// TIA Portal project "Mawomat" (V17)

(* hardware
DEVICE "S7-1500/ET200MP station_1"  S7-1500 station
   slot 0: "Rail_0"  Rack  6ES7 590-1***0-0AA0
   slot 1: "PLC_1"  CPU 1511-1 PN  6ES7 511-1AK00-0AB0  V1.8
      slot 3: "CPU display_1"  6ES7591-1AA00-0AA0
      slot 32768: "PROFINET interface_1"  X1
         slot 32769: "Port_1"  X1 P1
         slot 32770: "Port_2"  X1 P2
DEVICE "HMI_1"  KTP1200 Basic PN
   slot 0: "HMI_1"  KTP1200 Basic PN  6AV2 123-2MB03-0AX0  17.0.0.0
   slot 1: "HMI_RT_1"  KTP1200 Basic PN  6AV2 123-2MB03-0AX0  17.0.0.0
   slot 5: "HMI_1.IE_CP_1"  PROFINET Interface  17.0.0.0
      slot 1: "PROFINET Interface_1"  PROFINET Interface
         slot 1: "Port_1"  Port
DEVICE "SINAMICS G_1"  Sinamics.Device
   slot 0: "	_0"  Rail  SinamicsG120RackPN
   slot 0: "Drive_1"  G120 CU240E-2 PN  6SL3244-0BB12-1FA0  4.7.13
      slot 1: "PROFINET interface"  MDD-SinamicsG120-P
DEVICE "SINAMICS G_2"  Sinamics.Device
   slot 0: "	_0"  Rail  SinamicsG120RackPN
   slot 0: "Drive_2"  G120 CU240E-2 PN  6SL3244-0BB12-1FA0  4.7.13
      slot 1: "PROFINET interface"  MDD-SinamicsG120-P
*)

// ===== PLC "PLC_1"  CPU 1511-1 PN =====

VAR_GLOBAL   // PLC tag table "Default tag table"
   "System_Byte" AT %MB1 : Byte;
   "FirstScan" AT %M1.0 : Bool;
   "DiagStatusUpdate" AT %M1.1 : Bool;
   "AlwaysTRUE" AT %M1.2 : Bool;
   "AlwaysFALSE" AT %M1.3 : Bool;
   "Clock_Byte" AT %MB0 : Byte;
   "Clock_10Hz" AT %M0.0 : Bool;
   "Clock_5Hz" AT %M0.1 : Bool;
   "Clock_2.5Hz" AT %M0.2 : Bool;
   "Clock_2Hz" AT %M0.3 : Bool;
   "Clock_1.25Hz" AT %M0.4 : Bool;
   "Clock_1Hz" AT %M0.5 : Bool;
   "Clock_0.625Hz" AT %M0.6 : Bool;
   "Clock_0.5Hz" AT %M0.7 : Bool;
   "systemowe01" AT %M50.0 : Bool;
   "systemowe02" AT %M50.1 : Bool;
   "imp1s" AT %M50.2 : Bool;
   "Tag_29" AT %M51.0 : Bool;
   "Tag_28" AT %M51.1 : Bool;
   "imp0.1s" AT %M51.2 : Bool;
   "Tag_31" AT %M52.0 : Bool;
   "Tag_32" AT %M52.1 : Bool;
   "Imp0.2s" AT %M52.2 : Bool;
   "Tag_1" AT %M60.0 : Bool;
   "Tag_2" AT %M20.2 : Bool;
   "Tag_3" AT %M60.1 : Bool;
   "Tag_4" AT %M10.0 : Bool;
   "Tag_5" AT %M10.1 : Bool;
   "Tag_6" AT %M10.2 : Bool;
   "Tag_7" AT %M10.3 : Bool;
END_VAR

VAR_GLOBAL   // PLC tag table "Tag table_1"
   "qw256" AT %QW256 : Word;
END_VAR

TYPE "UDT321_DIO"
   STRUCT
      yNrPLC : Byte;   // DANE OGOLNE - Numer sterownika [0-255]
      yNrMAN : Byte;   // DANE OGOLNE - Numer powiazanej 'grupy recznej' [0-255]
      yNrID : Int;   // DANE OGOLNE - Numer ID obiektu w klasie [0-65536]
      yNrMD : Int;   // DANE OGOLNE - Numer powiazanego 'modelu drogi'
      bWeAkt : Bool;   // WEJSCIE - Aktywacja urz. w systemie (ustawiany tylko z programu)
      bWeZalAuto : Bool;   // WEJSCIE - Sterowanie urz. binarne w tr. Zdalnym-Auto: (0)- Wylacz; (1)- Zalacz
      bWeAwrZ : Bool;   // WEJSCIE - Awaria zewnetrzna: (0)-Brak; (1)-Aktywna
      bWeBlZmAuto : Bool;   // WEJŚCIE - Blokada zmiany trybu zdalnego z Auto na Man: (0)- Brak; (1)- Aktywna
      bRoZB1 : Byte := 16#5;   // !Rozkazy operetara
      bRoZB2 : Byte;   // !Rozkazy operatora - impulsy
      bSym : Word;   // !Symulacja
      bSt_Tryb : Word;   // !Stan
      bSt_Urz : Int;   // !Stan2
      bTrP : Int;   // !Tryb pracy
      bWySter : Bool;   // WYJSCIE - Sygnal zalaczenia urzadzenia
      bWyRst : Bool;   // WYJSCIE - Sygnal resetu awarii (impuls)
      yCzZadOpzZal : DWord;   // PARAMETR- Zadany czas opoznienia zalaczenia [0-255] sek.
      yCzAktOpzZal : DWord;   // PARAMETR- Aktualny czas opoznienia zalaczenia [0-255] sek.
      yCzZadOpzWyl : DWord;   // PARAMETR- Zadany czas opoznienia wylaczenia [0-255] sek.
      yCzAktOpzWyl : DWord;   // PARAMETR- Aktualny czas opoznienia wylaczenia [0-255] sek.
      bLatch : Bool;   // PARAMETR - Zatrzaskiwanie wyjscia (0) - Wylaczone; (1)-Zalaczone
      bAoff : Bool := 1;   // PARAMETR - samowylaczanie wylaczone (0); zalaczone (1)
      bHlp187 : Bool;   // WYJSCIE - Zal urz. w trybie AUTO
      bWeTrRem : Bool;
      bWeTrLok : Bool;
      bHlp186 : Bool;
      bTmr_On_Start : Bool;   // PARAMETR - Czas zadany timera filtru HH
      bTmr_Off_Start : Bool;   // PARAMETR - Czas zadany timera filtru LL
      bTmr_On_Ok : Bool;   // PARAMETR - Timer HH opoznienia zalaczenia odliczyl
      bTmr_Off_Ok : Bool;   // PARAMETR - Timer LL opoznienia zalaczenia odliczyl
   END_STRUCT;
END_TYPE

TYPE "UDT331_AI"
   STRUCT
      yNrPLC : Byte;   // DANE OGOLNE - Numer sterownika [0-255]
      yNrMAN : Byte;   // DANE OGOLNE - Numer powiazanej 'grupy recznej' [0-255]
      yNrID : Int;   // DANE OGOLNE - Numer ID obiektu w klasie [0-65536]
      yNrMD : Int;   // DANE OGOLNE - Numer powiazanego 'modelu drogi'
      bWeAkt : Bool;   // WEJSCIE - Aktywacja urz. w systemie (ustawiany tylko z programu)
      bWeAwrZ : Bool;   // WEJSCIE - Awaria zewnetrzna: (0)-Brak; (1)-Aktywna
      bWeBlZmAuto : Bool;   // WEJSCIE - Blokada zmiany trybu zdalnego z Auto na Man: (0)- Brak; (1)- Aktywna
      bWeSymUp : Bool;   // WEJSCIE - W trybie symulacji pomiaru skok w gore o rSymUp / sekunde
      bWeSymDown : Bool;   // WEJSCIE - W trybie symulacji pomiaru skok w dol o rSymDown / sekunde
      bRoZB1 : Byte := 16#01;   // !Rozkazy operetara
      bRoZB2 : Byte;   // !Rozkazy operatora - impulsy
      bSym : Word;   // !Symulacja
      bSt_Tryb : Word;   // !Stan
      bSt_Urz : Int;   // !Stan2
      bTrP : Int;   // !Tryb pracy
      bWyRst : Bool;   // WYJSCIE - Sygnal resetu awarii (impuls)
      yJednostka : Byte := 16#3;   // PARAMETR - Jednostka fizyczna
      yCzZadFiltru : Byte;   // PARAMETR - Czas zadany filtrow HH i LL [0-255] sek
      yCzasAktFiltrG : Byte := 16#3;   // PARAMETR - Czas aktualny filtru HH [0-255] sek
      yCzasAktFiltrD : Byte;   // PARAMETR - Czas aktualny filtru LL [0-255] sek
      bB : Byte;   // PARAMETR - Blokada generowania alarmow
      bAwrUst : Bool;   // PARAMETR - Reakcja na awarie toru pomiarowego: 0-na wyjsciu ZL; 1-ZH
      rZH : Real;   // PARAMETR - Zakres gorny pomiaru w jednostkach fizycznych
      rZL : Real;   // PARAMETR - Zakres dolny pomiaru w jednostkach fizycznych
      rGHH : Real;   // PARAMETR - Wartosc gornej granicy alarmowej w jednostkach fizycznych
      rGH : Real;   // PARAMETR - Wartosc gornej granicy ostrzegawczej w jednostkach fizycznych
      rGL : Real;   // PARAMETR - Wartosc dolnej granicy ostrzegawczej w jednostkach fizycznych
      rGLL : Real;   // PARAMETR - Wartosc gornej granicy alarmowej w jednostkach fizycznych
      rOffset : Real;   // PARAMETR - Offset pomiaru
      rFac : Real := 1.0;   // PARAMETR - Wspolczynnik skalujacy
      rSymUp : Real;   // PARAMETR - Wartosc zmiany w gore w czasie 1sek. w trybie symulacji pomiaru
      rSymDown : Real;   // PARAMETR - Wartosc zmiany w dol w czasie 1 sek. w trybie symulacji pomiaru
      wWe : Word;   // WEJSCIE - Sygnal z wejscia PIW
      rRoManSter : Real;   // ROZKAZ OPERATORA - wartosc pomiaru wpisana w trybie Zdalnym-Recznym
      rWy : Real;   // WYJSCIE - Syngal wyjsciowy pomiaru w jednostkach fizycznych
      yWy : Int := 16#3;   // WYJSCIE - Sygnal wyjsciowy pomiaru (0-100%)
      dTmr_HH_Start : Bool;   // PARAMETR - Czas zadany timera filtru HH
      dTmr_LL_Start : Bool;   // PARAMETR - Czas zadany timera filtru LL
      dTmr_HH_Ok : Bool;   // PARAMETR - Timer HH opoznienia zalaczenia odliczyl
      dTmr_LL_Ok : Bool;   // PARAMETR - Timer LL opoznienia zalaczenia odliczyl
   END_STRUCT;
END_TYPE

TYPE "UDT322_DVI"
   STRUCT
      yNrPLC : Byte;   // DANE OGOLNE - Numer sterownika [0-255]
      yNrMAN : Byte;   // DANE OGOLNE - Numer powiazanej 'grupy recznej' [0-255]
      yNrID : Int;   // DANE OGOLNE - Numer ID obiektu w klasie [0-65536]
      yNrMD : Int;   // DANE OGOLNE - Numer powiazanego 'modelu drogi'
      bWeAkt : Bool;   // WEJSCIE - Aktywacja urz. w systemie (ustawiany tylko z programu)
      bWeZalAuto : Bool;   // WEJSCIE - Sterowanie urz. binarne w tr. Zdalnym-Auto: (0)- Wylacz; (1)- Zalacz
      bWePotwZal : Bool;   // WEJSCIE - Potwiedzenie zalaczenia/otwarcia
      bWePotwWyl : Bool;   // WEJSCIE - Potwierdzenie wylaczenia/zamkniecia
      bWePotwGot : Bool;   // WEJSCIE - Potwierdzenie gotowosci
      bWeTrLok : Bool;   // WEJSCIE - Tryb sterowania: 0-Zdalne z PC; 1-Lokalne z elewacji szafy
      bWeTrRem : Bool;   // WEJSCIE - Tryb remontowy (z wylacznika): 0-Brak; 1-Aktywny
      bWeAwrZ : Bool;   // WEJSCIE - Awaria zewnetrzna: (0)-Brak; (1)-Aktywna
      bWeBlZmAuto : Bool;   // WEJŚCIE - Blokada zmiany trybu zdalnego z Auto na Man: (0)- Brak; (1)- Aktywna
      bWeIlock : Bool;   // WEJSCIE - Interlock w trybie Zdalnym-Auto: 0-Brak; 1-Aktywny
      bRoZB1 : Byte := 16#01;   // !Rozkazy operetara
      bRoZB2 : Byte;   // !Rozkazy operatora - impulsy
      bSym : Word;   // !Symulacja
      bSt_Tryb : Word;   // !Stan
      bSt_Urz : Int;   // !Stan2
      bTrP : Int;   // !Tryb pracy
      bWySter : Bool;   // WYJSCIE - Sygnal zalaczenia urzadzenia
      bWyRst : Bool;   // WYJSCIE - Sygnal resetu awarii (impuls)
      yCzZadOpzZal : DWord;   // PARAMETR- Zadany czas opoznienia zalaczenia [0-255] sek.
      yCzAktOpzZal : DWord;   // PARAMETR- Aktualny czas opoznienia zalaczenia [0-255] sek.
      yCzZadOpzWyl : DWord;   // PARAMETR- Zadany czas opoznienia wylaczenia [0-255] sek.
      yCzAktOpzWyl : DWord;   // PARAMETR- Aktualny czas opoznienia wylaczenia [0-255] sek.
      yCzZadOpzAlm : Byte;   // PARAMETR - Zadany czas opoznienia alarmu od potwierdzen [0-255] sek
      yCzasAktOpzAlm : Byte;   // PARAMETR - Aktualny czas opoznienia alarmu od potwierdzen [0-255] sek
      bNoNc : Bool;   // PARAMETR - Zawor NC-0; Zawor NO-1
      bAoff : Bool := 1;   // PARAMETR - samowylaczanie wylaczone (0); zalaczone (1)
      bTmr_On_Start : Bool;   // PARAMETR - Sygnal startu timera zalaczenia urzadzenia
      bTmr_Off_Start : Bool;   // PARAMETR - Sygnal startu timera wylaczenia urzadzenia
      bTmr_Awr_Start : Bool;   // PARAMETR - Sygnal startu timera awarii urzadzenia
      bTmr_On_Ok : Bool;   // PARAMETR - Sygnal odliczenia czasu zalaczenia urz.
      bTmr_Off_Ok : Bool;   // PARAMETR - Sygnal odliczenia czasu wylaczenia urz.
      bTmr_Alm_Ok : Bool;   // PARAMETR - Sygnal odliczenia czasu awarii urz.
      bHlp184 : Bool;
      bHlp185 : Bool;
      bHlp186 : Bool;
      bHlp187 : Bool;
      bHlp256 : Bool;
      bHlp257 : Bool;
      bHlp_NoNc : Bool;   // 1- zawsze otwieranie; 0-zawsze zamykanie
   END_STRUCT;
END_TYPE

TYPE "UDT323_DM1"
   STRUCT
      yNrPLC : Byte;   // DANE OGOLNE - Numer sterownika [0-255]
      yNrMAN : Byte;   // DANE OGOLNE - Numer powiazanej 'grupy recznej' [0-255]
      yNrID : Int;   // DANE OGOLNE - Numer ID obiektu w klasie [0-65536]
      yNrMD : Int;   // DANE OGOLNE - Numer powiazanego 'modelu drogi'
      bWeAkt : Bool;   // WEJSCIE - Aktywacja urz. w systemie (ustawiany tylko z programu)
      bWeZalAuto : Bool;   // WEJSCIE - Sterowanie urz. binarne w tr. Zdalnym-Auto: (0)- Wylacz; (1)- Zalacz
      bWePotwZal : Bool;   // WEJSCIE - Potwiedzenie zalaczenia/otwarcia
      bWePotwWyl : Bool;   // WEJSCIE - Potwierdzenie wylaczenia/zamkniecia
      bWePotwGot : Bool;   // WEJSCIE - Potwierdzenie gotowosci
      bWeTrLok : Bool;   // WEJSCIE - Tryb sterowania: 0-Zdalne z PC; 1-Lokalne z elewacji szafy
      bWeTrRem : Bool;   // WEJSCIE - Tryb remontowy (z wylacznika): 0-Brak; 1-Aktywny
      bWeAwrZ : Bool;   // WEJSCIE - Awaria zewnetrzna: (0)-Brak; (1)-Aktywna
      bWeBlZmAuto : Bool;   // WEJSCIE - Blokada zmiany trybu zdalnego z Auto na Man: (0)- Brak; (1)- Aktywna
      bWeIlock : Bool;   // WEJSCIE - Interlock w trybie Zdalnym-Auto: 0-Brak; 1-Aktywny
      bWeKier : Bool;   // WEJSCIE - Kierunek obrotow: 0-Prawo; 1-Lewo
      bRoZB1 : Byte := 16#01;   // !Rozkazy operetara
      bRoZB2 : Byte;   // !Rozkazy operatora - impulsy
      bSym : Word;   // !Symulacja
      bSt_Tryb : Word;   // !Stan
      bSt_Urz : Int;   // !Stan2
      bTrP : Int;   // !Tryb pracy
      bWySter : Bool;   // WYJSCIE - Sygnal zalaczenia urzadzenia
      bWyRst : Bool;   // WYJSCIE - Sygnal resetu awarii (impuls)
      bWyKier : Bool;   // WYJSCIE - Sygnal kierunku obrotow: 0-Prawo; 1-Lewo
      yCzZadOpzZal : DWord;   // PARAMETR- Zadany czas opoznienia zalaczenia [0-255] sek.
      yCzAktOpzZal : DWord;   // PARAMETR- Aktualny czas opoznienia zalaczenia [0-255] sek.
      yCzZadOpzWyl : DWord;   // PARAMETR- Zadany czas opoznienia wylaczenia [0-255] sek.
      yCzAktOpzWyl : DWord;   // PARAMETR- Aktualny czas opoznienia wylaczenia [0-255] sek.
      yCzZadOpzAlm : Byte;   // PARAMETR - Zadany czas opoznienia alarmu od potwierdzen [0-255] sek
      yCzasAktOpzAlm : Byte;   // PARAMETR - Aktualny czas opoznienia alarmu od potwierdzen [0-255] sek
      bKier : Bool;   // PARAMETR - Bit wyboru stacyjki (tylko z wejscia bloku logiki)
      bAoff : Bool := 1;   // PARAMETR - samowylaczanie wylaczone (0); zalaczone (1)
      bTmr_On_Start : Bool;   // PARAMETR - Sygnal startu timera zalaczenia urzadzenia
      bTmr_Off_Start : Bool;   // PARAMETR - Sygnal startu timera wylaczenia urzadzenia
      bTmr_Awr_Start : Bool;   // PARAMETR - Sygnal startu timera awarii urzadzenia
      bTmr_On_Ok : Bool;   // PARAMETR - Sygnal odliczenia czasu zalaczenia urz.
      bTmr_Off_Ok : Bool;   // PARAMETR - Sygnal odliczenia czasu wylaczenia urz.
      bTmr_Alm_Ok : Bool;   // PARAMETR - Sygnal odliczenia czasu awarii urz.
      bHlp186 : Bool;
      bHlp187 : Bool;
      bHlp256 : Bool := false;
      bHlp257 : Bool;
   END_STRUCT;
END_TYPE

TYPE "UDT332_AO"
   STRUCT
      yNrPLC : Byte;   // DANE OGOLNE - Numer sterownika [0-255]
      yNrMAN : Byte;   // DANE OGOLNE - Numer powiazanej 'grupy recznej' [0-255]
      yNrID : Int;   // DANE OGOLNE - Numer ID obiektu w klasie [0-65536]
      yNrMD : Int;   // DANE OGOLNE - Numer powiazanego 'modelu drogi'
      bWeAkt : Bool;   // WEJSCIE - Aktywacja urz. w systemie (ustawiany tylko z programu)
      bWeAwrZ : Bool;   // WEJSCIE - Awaria zewnetrzna: (0)-Brak; (1)-Aktywna
      bWeBlZmAuto : Bool;   // WEJSCIE - Blokada zmiany trybu zdalnego z Auto na Man: (0)- Brak; (1)- Aktywna
      bRoZB1 : Byte := 16#01;   // !Rozkazy operetara
      bRoZB2 : Byte;   // !Rozkazy operatora - impulsy
      bSym : Word;   // !Symulacja
      bSt_Tryb : Word;   // !Stan
      bSt_Urz : Int;   // !Stan2
      bTrP : Int;   // !Tryb pracy
      bWyRst : Bool;   // WYJSCIE - Sygnal resetu awarii (impuls)
      yJednostka : Byte := 16#3;   // PARAMETR - Jednostka fizyczna
      yCzZadFiltru : Byte;   // PARAMETR - Czas zadany filtrow HH i LL [0-255] sek
      yCzasAktFiltrG : Byte := 16#3;   // PARAMETR - Czas aktualny filtru HH [0-255] sek
      yCzasAktFiltrD : Byte;   // PARAMETR - Czas aktualny filtru LL [0-255] sek
      bB : Byte;   // PARAMETR - Blokada generowania alarmow
      bAwrUst : Bool;   // PARAMETR - Reakcja na awarie toru pomiarowego: 0-na wyjsciu ZL; 1-ZH
      rZH : Real;   // PARAMETR - Zakres gorny pomiaru w jednostkach fizycznych
      rZL : Real;   // PARAMETR - Zakres dolny pomiaru w jednostkach fizycznych
      rGHH : Real;   // PARAMETR - Wartosc gornej granicy alarmowej w jednostkach fizycznych
      rGH : Real;   // PARAMETR - Wartosc gornej granicy ostrzegawczej w jednostkach fizycznych
      rGL : Real;   // PARAMETR - Wartosc dolnej granicy ostrzegawczej w jednostkach fizycznych
      rGLL : Real;   // PARAMETR - Wartosc gornej granicy alarmowej w jednostkach fizycznych
      rOffset : Real;   // PARAMETR - Offset pomiaru
      rFac : Real := 1.0;   // PARAMETR - Wspolczynnik skalujacy
      rHI_LIM : Real;   // PARAMETR - Zakres gorny wielkosci fizycznej
      rWe : Real;   // WEJSCIE - Sygnal z wejscia programu
      rRoManSter : Real;   // ROZKAZ OPERATORA - wartosc pomiaru wpisana w trybie Zdalnym-Recznym
      wWy : Word;   // WYJSCIE - Sygnal na wyjscie PQW/QW
      rWy : Real;   // WYJSCIE - Syngal wyjsciowy pomiaru w real
      yWy : Byte := 16#3;   // WYJSCIE - Sygnal wyjsciowy pomiaru (0-100%)
      dTmr_HH_Start : Bool;   // PARAMETR - Czas zadany timera filtru HH
      dTmr_LL_Start : Bool;   // PARAMETR - Czas zadany timera filtru LL
      dTmr_HH_Ok : Bool;   // PARAMETR - Timer HH opoznienia zalaczenia odliczyl
      dTmr_LL_Ok : Bool;   // PARAMETR - Timer LL opoznienia zalaczenia odliczyl
   END_STRUCT;
END_TYPE

TYPE "UDT352_FF8"
   STRUCT
      yNrPLC : Byte;   // DANE OGOLNE - Numer sterownika [0-255]
      yNrMAN : Byte;   // DANE OGOLNE - Numer powiazanej 'grupy recznej' [0-255]
      yNrID : Int;   // DANE OGOLNE - Numer ID obiektu w klasie [0-65536]
      yNrMD : Int;   // DANE OGOLNE - Numer powiazanego 'modelu drogi'
      bWeAkt : Bool;   // WEJSCIE - Aktywacja urz. w systemie (ustawiany tylko z programu)
      bWeZalAuto : Bool;   // WEJSCIE - Sterowanie urz. binarne w tr. Zdalnym-Auto: (0)- Wylacz; (1)- Zalacz
      bWeBlZmAuto : Bool;   // WEJSCIE - Blokada zmiany trybu zdalnego z Auto na Man: (0)- Brak; (1)- Aktywna
      bWeIlock : Bool;   // WEJSCIE - Interlock w trybie Zdalnym-Auto: 0-Brak; 1-Auto
      bWeZeruj : Bool;   // WEJSCIE - Zerowanie timera (kasowanie przez obiekt)
      bRoZB1 : Byte := 16#01;   // !Rozkazy operetara
      bSym : Word;   // !Symulacja
      bSt_Tryb : Word;   // !Stan
      bSt_Urz : Int;   // !Stan2
      bTrP : Int;   // !Tryb pracy
      bWySter : Bool;   // WYJSCIE - Sygnal zalaczenia urzadzenia
      yJednostka : Byte;   // PARAMETR - Jednostka zliczania czasu
      bIhlp : Bool;   // Pomocnicze sterowanie impulsem
      bPauza : Bool;   // Bit pauzy miedzy grupami impulsow
      bI1 : Bool;   // Wyjscie dla impulsu 1
      bI2 : Bool;   // Wyjscie dla impulsu 2
      bI3 : Bool;   // Wyjscie dla impulsu 3
      bI4 : Bool;   // Wyjscie dla impulsu 4
      bI5 : Bool;   // Wyjscie dla impulsu 5
      bI6 : Bool;   // Wyjscie dla impulsu 6
      bI7 : Bool;   // Wyjscie dla impulsu 7
      bI8 : Bool;   // Wyjscie dla impulsu 8
      bAoff : Bool;   // PARAMETR - samowylacznie: 0-wylaczone; 1-zalaczone
      iIG : Int;   // Ilosc grup
      dT1_old : DInt;   // Zadany czas impulsu
      dT2 : DInt;   // Zadany czas przerwy miedzy impulsami
      dT3 : DInt;   // Zadany czas przerwy miedzy grupami impulsow
      dT1_Akt : DInt;   // Aktualny czas impulsu
      dT2_Akt : DInt := 0;   // Aktualny czas przerwy miedzy impulsami
      dT3_Akt : DInt := 0;   // Aktualny czas przerwy miedzy grupami impulsow
      iPetle : Int;   // Licznik impulsow (zakonczonych)
      dT1i : DInt;   // Zadany czas impulsu 1
      dT2i : DInt;   // Zadany czas impulsu 2
      dT3i : DInt;   // Zadany czas impulsu 3
      dT4i : DInt;   // Zadany czas impulsu 4
      dT5i : DInt;   // Zadany czas impulsu 5
      dT6i : DInt;   // Zadany czas impulsu 6
      dT7i : DInt;   // Zadany czas impulsu 7
      dT8i : DInt;   // Zadany czas impulsu 8
      dwBlokSCADA : DWord;   // Blokada parametrow na SCADA
   END_STRUCT;
END_TYPE

TYPE "UDT340_PID"
   STRUCT
      yNrPLC : Byte;   // DANE OGOLNE - Numer sterownika [0-255]
      yNrMAN : Byte;   // DANE OGOLNE - Numer powiazanej 'grupy recznej' [0-255]
      yNrID : Int;   // DANE OGOLNE - Numer ID obiektu w klasie [0-65536]
      yNrMD : Int;   // DANE OGOLNE - Numer powiazanego 'modelu drogi'
      bWeAkt : Bool;   // WEJSCIE - Aktywacja urz. w systemie (ustawiany tylko z programu)
      bWeZalAuto : Bool;   // WEJSCIE - Sterowanie urz. binarne w tr. Zdalnym-Auto: (0)- Wylacz; (1)- Zalacz
      bWeBlZmAuto : Bool;   // WEJSCIE - Blokada zmiany trybu zdalnego z Auto na Man: (0)- Brak; (1)- Aktywna
      bWeTrck : Bool;   // WEJSCIE - Sledzenie: 0-Wylaczone; 1-Zalaczone
      bRoZB1 : Byte := 16#01;   // !Rozkazy operetara
      bSym : Word;   // !Symulacja
      bSt_Tryb : Word;   // !Stan
      bSt_Urz : Int;   // !Stan2
      bTrP : Int;   // !Tryb pracy
      bWySter : Bool;   // WYJSCIE - Sygnal zalaczenia urzadzenia
      QLMN_HLM : Bool;   // WYJSCIE -
      QLMN_LLM : Bool;   // WYJSCIE -
      sbArwHLmOn : Bool;   // WYJSCIE -
      sbArwLLmOn : Bool;   // WYJSCIE -
      bHlp187 : Bool;   // Bit pomocniczy On/Off
      yJednostka : Byte := 16#3;   // PARAMETR - Jednostka fizyczna
      rTrace : Real;   // PARAMETR - Wartosc wejsciowa dla sygnalu sledzenia (0-100%)
      PVPER_ON : Bool;   // PARAMETR -
      P_SEL : Bool := true;   // PARAMETR -
      I_SEL : Bool;   // PARAMETR -
      INT_HOLD : Bool;   // PARAMETR -
      I_ITL_ON : Bool;   // PARAMETR -
      D_SEL : Bool;   // PARAMETR -
      bAoff : Bool;   // PARAMETR -
      CYCLE : Real := 0.1;   // PARAMETR -
      SP_INT : Real;   // PARAMETR -
      PV_IN : Real;   // PARAMETR -
      PV_PER : Word;   // PARAMETR -
      MAN : Real;   // PARAMETR -
      GAIN : Real := 2.0;   // PARAMETR -
      TI : Real := 1.0;   // PARAMETR -
      TD : Real;   // PARAMETR -
      TM_LAG : Real;   // PARAMETR -
      DEADB_W : Real;   // PARAMETR -
      LMN_HLM : Real := 1.0;   // PARAMETR -
      LMN_LLM : Real;   // PARAMETR -
      PV_FAC : Real := 1.0;   // PARAMETR -
      PV_OFF : Real;   // PARAMETR -
      LMN_FAC : Real := 1.0;   // PARAMETR -
      LMN_OFF : Real;   // PARAMETR -
      I_ITLVAL : Real;   // PARAMETR -
      DISV : Real;   // PARAMETR -
      LMN : Real;   // PARAMETR -
      LMN_PER : Word;   // PARAMETR -
      LMN_P : Real;   // PARAMETR -
      LMN_I : Real;   // PARAMETR -
      LMN_D : Real;   // PARAMETR -
      PV : Real;   // PARAMETR -
      ER : Real;   // PARAMETR -
      sinvAlt : Real;   // PARAMETR -
      sIanteilAlt : Real;   // PARAMETR -
      sRestInt : Real;   // PARAMETR -
      sRestDif : Real;   // PARAMETR -
      sRueck : Real;   // PARAMETR -
      sRueckOld : Real;   // PARAMETR -
      sLmn : Real;   // PARAMETR -
      ErKp : Real;   // PARAMETR - Uchyb regulacji
      Ianteil : Real;   // TEMP
      Panteil : Real;   // TEMP
      Danteil : Real;   // TEMP
      Diff : Real;   // TEMP
      "L78.2" : Bool;   // TEMP
      dLmn : Real;
      rVal : Real;
   END_STRUCT;
END_TYPE

TYPE "UDT350_Sek"
   STRUCT
      yNrMan : Byte;   // Numer powiazanego obiektu Man
      bAkt : Bool := 1;   // Bit aktywacji obiektu. 1- obiekt aktywowany; 0-obiekt nieaktywowany
      bSe_ReqStart : Bool;   // ROZKAZ - Start sekwencji
      bSe_ReqStop : Bool;   // ROZKAZ - Stop sekwencji
      bSe_ReqPauza : Bool;   // ROZKAZ - Pauza sekwencji
      bSe_ReqWznow : Bool;   // ROZKAZ - Wznowienie po pauzie sekwencji
      bSe_ReqRestart : Bool;   // ROZKAZ - Restart sekwencji
      bSe_ReqZmiana : Bool;   // ROZKAZ (wewnetrzny) - Zmiana kroku sekwencji
      bSe_Hlp1 : Bool;   // Bit pomocniczy
      bSe_Wylaczony : Bool;   // STAN - Sekwencja wylaczona
      bSe_Run : Bool;   // STAN - Sekwencja zalaczona
      bSe_Pauza : Bool;   // STAN - Sekwencja w pauzie
      bSe_Interlok : Bool;   // STAN - Sekwencja w blokadzie startu
      ySe_NrKrokSel : Byte := 16#1;   // STAN - Numer aktualnie uzywanego kroku
      ySe_MaxKrok : Byte := 16#1;   // STAN - Ilosc dostepnych krokow
      Rez : Array[1..10] of Byte;
      Krok : Array[1..96] of Struct
         bRun : Bool;   // STAN - Krok xxx Run
         bPauza : Bool;   // STAN - Krok xxx Pauza
         bHlp1 : Bool;
         bHlp2 : Bool;
         bHlp3 : Bool;
         bHlp4 : Bool;
         bW1 : Bool;   // ROZKAZ - warunek przejscia do korku #bKrokxxx_NastW1
         bW2 : Bool;   // ROZKAZ - warunek przejscia do korku #bKrokxxx_NastW2
         yNastW1 : Byte;   // Numer kroku do ktorego skaczemy przy ust. #bKrokxxx_NastW1
         yNastW2 : Byte;   // Numer kroku do ktorego skaczemy przy ust. #bKrokxxx_NastW2
         yAlarm : Byte;
      END_STRUCT;
   END_STRUCT;
END_TYPE

TYPE "LSim_typeZone"
// V1.1
   STRUCT
      inputHeat : Real;   // input value in REAL format - heating / Ausgangswert im REAL-Format - Heizen
      inputCool : Real;   // input value in REAL format - cooling / Ausgangswert im REAL-Format - Kühlen
      disturbance : Real;   // disturbance (input)
      output : Real;   // zone temperature (output)
   END_STRUCT;
END_TYPE

TYPE "UDT353_TMR"
   STRUCT
      yNrPLC : Byte;   // DANE OGOLNE - Numer sterownika [0-255]
      yNrMAN : Byte;   // DANE OGOLNE - Numer powiazanej 'grupy recznej' [0-255]
      yNrID : Int;   // DANE OGOLNE - Numer ID obiektu w klasie [0-65536]
      yNrMD : Int;   // DANE OGOLNE - Numer powiazanego 'modelu drogi'
      bWeAkt : Bool;   // WEJSCIE - Aktywacja urz. w systemie (ustawiany tylko z programu)
      bWeZalAuto : Bool;   // WEJSCIE - Sterowanie urz. binarne w tr. Zdalnym-Auto: (0)- Wylacz; (1)- Zalacz
      bWeBlZmAuto : Bool;   // WEJSCIE - Blokada zmiany trybu zdalnego z Auto na Man: (0)- Brak; (1)- Aktywna
      bWeIlock : Bool;   // WEJSCIE - Interlock w trybie Zdalnym-Auto: 0-Brak; 1-Auto
      bWeZeruj : Bool;   // WEJSCIE - Zerowanie timera (kasowanie przez obiekt)
      bRoZB1 : Byte := 16#01;   // !Rozkazy operetara
      bSym : Word;   // !Symulacja
      bSt_Tryb : Word;   // !Stan
      bSt_Urz : Int;   // !Stan2
      bTrP : Int;   // !Tryb pracy
      bWySter : Bool;   // WYJSCIE - Sygnal zalaczenia urzadzenia
      bHlp187 : Bool;
      yJednostka : Byte;   // PARAMETR - Jednostka zliczania czasu
      dCzZad : DWord;   // PARAMETR - Zadany czas [sek].
      bLatch : Bool;   // PARAMETR - Zamrozenie wyjsc: 0- wylaczone; 1- zalaczone
      bAoff : Bool := 1;   // PARAMETR - samowylaczanie wylaczone: 0-wylaczone; 1- zalaczone
      dCzAkt : DWord;   // PARAMETR - Aktualny czas [sek].
   END_STRUCT;
END_TYPE

TYPE "LSim_typeDynState"
// V1.1
   STRUCT
      kInt : Real := 0.2;   // coupling constant internal
      kFor : Real := 0.3;   // coupling constant forwards
      kBack : Real := 0.1;   // coupling constant backwards
      uInp : Real;   // uInp = heatPT1out - coolPT1out + disturbance
      u : Real;   // u = uInp + kFor(z-1) * y(z-1) - 2 * kInt * y + kBack(z+1) * y(z+1); z = zone
      y : Real;   // y = PT2out
   END_STRUCT;
END_TYPE

DATA_BLOCK "Sequences_DB"   // DB4
{ S7_Optimized_Access := 'TRUE' }
VERSION : 0.1
// stored: InstanceOfName Sequence1
"Sequence1"
BEGIN
END_DATA_BLOCK

// folder: DI

DATA_BLOCK "DI_Objects_DB"   // DB10
{ S7_Optimized_Access := 'TRUE' }
VERSION : 0.1
// stored: InstanceOfName DI_Objects
"DI_Objects"
BEGIN
END_DATA_BLOCK

// folder: DV

DATA_BLOCK "DV_Objects_DB"   // DB11
{ S7_Optimized_Access := 'TRUE' }
VERSION : 0.1
// stored: InstanceOfName DV_Objects
"DV_Objects"
BEGIN
END_DATA_BLOCK

// folder: LSim

DATA_BLOCK "LSim_PT3_DB"   // DB9
{ S7_Optimized_Access := 'TRUE' }
VERSION : 2.01
// stored: InstanceOfName LSim_PT3
"LSim_PT3"
BEGIN
END_DATA_BLOCK

// folder: Mawomat_stare/Klasy_DB

DATA_BLOCK "DB321_DIO"   // DB321
{ S7_Optimized_Access := 'TRUE' }
VERSION : 0.1
   VAR RETAIN
      DIO : Array[1..150] of "UDT321_DIO";
   END_VAR
BEGIN
END_DATA_BLOCK

DATA_BLOCK "DB322_DV1"   // DB322
{ S7_Optimized_Access := 'TRUE' }
VERSION : 0.1
   VAR RETAIN
      DV1 : Array[1..4] of "UDT322_DVI";
   END_VAR
BEGIN
END_DATA_BLOCK

DATA_BLOCK "DB323_DM1"   // DB323
{ S7_Optimized_Access := 'TRUE' }
VERSION : 0.1
   VAR RETAIN
      DM1 : Array[1..30] of "UDT323_DM1";
   END_VAR
BEGIN
   DM1[2].bRoZB1 := 16#05;
   DM1[3].bRoZB1 := 16#05;
   DM1[4].bRoZB1 := 16#05;
   DM1[5].bRoZB1 := 16#05;
   DM1[6].bRoZB1 := 16#05;
   DM1[3].bWeAkt := true;
   DM1[2].bWeAkt := true;
   DM1[4].bWeAkt := true;
   // DM1[2] : Wozek glowny
   // DM1[3] : Wozek dodatkowy
   // DM1[4] : Wciagarka glowna silnik 1
   // DM1[5] : Wciagarka pomocnicza
   // DM1[6] : Chwytak
   // DM1[1] : Most
   // DM1[14] : Wciagarka glowna silnik 2
   // DM1[7] : Chwytak pomocniczy
END_DATA_BLOCK

DATA_BLOCK "DB331_AI"   // DB331
{ S7_Optimized_Access := 'TRUE' }
VERSION : 0.1
   VAR RETAIN
      AI : Array[1..10] of "UDT331_AI";
   END_VAR
BEGIN
   AI[1].rZH := 20.0;
   AI[1].rZL := 0.0;
   AI[1].rGHH := 7.1;
   AI[1].rGH := 4.5;
   AI[1].rGL := -1.0;
   AI[1].rGLL := -2.0;
   AI[1].rOffset := 0.1;
   AI[1].rFac := 0.1;
   AI[2].rZH := 20.0;
   AI[2].rZL := 0.0;
   AI[2].rGHH := 7.1;
   AI[2].rGH := 4.5;
   AI[2].rGL := -1.0;
   AI[2].rGLL := -2.0;
   AI[2].rOffset := 0.1;
   AI[2].rFac := 0.1;
   AI[3].rZH := 300.0;
   AI[3].rZL := 0.0;
   AI[3].rGHH := 300.0;
   AI[3].rGH := 300.0;
   AI[3].rGL := 50.0;
   AI[3].rGLL := 20.0;
   AI[3].rOffset := 1.0;
   AI[3].rFac := 1.0;
   AI[4].rZH := 0.0;
   AI[4].rZL := 0.0;
   AI[4].rGHH := 0.0;
   AI[4].rGH := 0.0;
   AI[4].rGL := 0.0;
   AI[4].rGLL := 0.0;
   AI[4].rOffset := 0.0;
   AI[4].rFac := 1.0;
   AI[5].rZH := 2764.8;
   AI[5].rZL := 0.0;
   AI[5].rGHH := 90.0;
   AI[5].rGH := 80.0;
   AI[5].rGL := 0.0;
   AI[5].rGLL := 0.0;
   AI[5].rOffset := 10.0;
   AI[5].rFac := 1.0;
   AI[6].rZH := 2764.8;
   AI[6].rZL := 0.0;
   AI[6].rGHH := 90.0;
   AI[6].rGH := 80.0;
   AI[6].rGL := 0.0;
   AI[6].rGLL := 0.0;
   AI[6].rOffset := 10.0;
   AI[6].rFac := 1.0;
   AI[7].rZH := 2764.8;
   AI[7].rZL := 0.0;
   AI[7].rGHH := 150.0;
   AI[7].rGH := 130.0;
   AI[7].rGL := 0.0;
   AI[7].rGLL := 0.0;
   AI[7].rOffset := 10.0;
   AI[7].rFac := 1.0;
   AI[8].rZH := 2764.8;
   AI[8].rZL := 0.0;
   AI[8].rGHH := 150.0;
   AI[8].rGH := 130.0;
   AI[8].rGL := 0.0;
   AI[8].rGLL := 0.0;
   AI[8].rOffset := 10.0;
   AI[8].rFac := 1.0;
   AI[9].rZH := 2764.8;
   AI[9].rZL := 0.0;
   AI[9].rGHH := 150.0;
   AI[9].rGH := 130.0;
   AI[9].rGL := 0.0;
   AI[9].rGLL := 0.0;
   AI[9].rOffset := 10.0;
   AI[9].rFac := 1.0;
   AI[10].rZH := 300.0;
   AI[10].rZL := 0.0;
   AI[10].rGHH := 0.0;
   AI[10].rGH := 0.0;
   AI[10].rGL := 50.0;
   AI[10].rGLL := 20.0;
   AI[10].rOffset := 10.0;
   AI[10].rFac := 1.0;
   // AI[1] : Main Drive - Vibration DE
   // AI[2] : Main Drive - Vibration NDE
   // AI[3] : Main Drive - Cooling Water Flow 2
   // AI[4] : Spare
   // AI[5] : Main Drive - Bearing Temp DE
   // AI[6] : Main Drive - Bearing Temp NDE
   // AI[7] : Main Drive - Winding U Temp
   // AI[8] : Main Drive - Winding V Temp
   // AI[9] : Main Drive - Winding W Temp
   // AI[10] : Main Drive - Cooling Water Flow Induction
END_DATA_BLOCK

DATA_BLOCK "DB332_AO"   // DB332
{ S7_Optimized_Access := 'TRUE' }
VERSION : 0.1
   VAR RETAIN
      AO : Array[1..10] of "UDT332_AO";
   END_VAR
BEGIN
END_DATA_BLOCK

DATA_BLOCK "DB340_PID"   // DB340
{ S7_Optimized_Access := 'TRUE' }
VERSION : 0.1
   VAR RETAIN
      PID : Array[1..5] of "UDT340_PID";
   END_VAR
BEGIN
END_DATA_BLOCK

DATA_BLOCK "DB350_SEK"   // DB350
{ S7_Optimized_Access := 'FALSE' }
VERSION : 0.1
   VAR
      SEK_Odwijak1_Otwieranie : "UDT350_Sek";
   END_VAR
BEGIN
END_DATA_BLOCK

DATA_BLOCK "DB352_FF8"   // DB352
{ S7_Optimized_Access := 'TRUE' }
VERSION : 0.1
   VAR RETAIN
      FF8 : Array[1..5] of "UDT352_FF8";
   END_VAR
BEGIN
END_DATA_BLOCK

DATA_BLOCK "DB353_TMR"   // DB353
{ S7_Optimized_Access := 'TRUE' }
VERSION : 0.1
   VAR
      TMR : Array[1..10] of "UDT353_TMR";
   END_VAR
BEGIN
END_DATA_BLOCK

// folder: Sinamics

DATA_BLOCK "DB_Sinamics"   // DB1
{ S7_Optimized_Access := 'TRUE' }
VERSION : 0.1
// stored: InstanceOfName DM_Sinamics
"DM_Sinamics"
BEGIN
END_DATA_BLOCK

DATA_BLOCK "DB_DM"   // DB2
{ S7_Optimized_Access := 'TRUE' }
VERSION : 0.1
// stored: InstanceOfName DM_Objects
"DM_Objects"
BEGIN
END_DATA_BLOCK

// folder: (top level)

DATA_BLOCK "pump2"   // DB3, Motion_DB
{ S7_Optimized_Access := 'TRUE' }
AUTHOR : SIMATIC
FAMILY : MC_1500
VERSION : 2.0
// stored: InstanceOfName TO_SpeedAxis
"TO_SpeedAxis"
BEGIN
   DynamicLimits.MaxAcceleration := 1000.0;
   DynamicLimits.MaxDeceleration := 1000.0;
   DynamicLimits.MaxJerk := 20000.0;
   DynamicDefaults.Acceleration := 200.0;
   DynamicDefaults.Deceleration := 200.0;
   DynamicDefaults.Jerk := 4000.0;
   DynamicDefaults.EmergencyDeceleration := 1000.0;
   Actor.Interface.AddressIn := 260;
   Actor.Interface.AddressOut := 260;
END_DATA_BLOCK

DATA_BLOCK "pump1"   // DB5, Motion_DB
{ S7_Optimized_Access := 'TRUE' }
AUTHOR : SIMATIC
FAMILY : MC_1500
VERSION : 2.0
// stored: InstanceOfName TO_SpeedAxis
"TO_SpeedAxis"
BEGIN
   DynamicLimits.MaxAcceleration := 1000.0;
   DynamicLimits.MaxDeceleration := 1000.0;
   DynamicLimits.MaxJerk := 20000.0;
   DynamicDefaults.Acceleration := 200.0;
   DynamicDefaults.Deceleration := 200.0;
   DynamicDefaults.Jerk := 4000.0;
   DynamicDefaults.EmergencyDeceleration := 1000.0;
   Actor.Interface.AddressIn := 256;
   Actor.Interface.AddressOut := 256;
   Simulation.Mode := 1;
END_DATA_BLOCK

FUNCTION_BLOCK "Sequencer"   // FB3, SCL
{ S7_Optimized_Access := 'TRUE' }
VERSION : 0.1
   VAR_INPUT
      inStart : Bool;
      inNexStepNb : Int;
      inManualMode : Bool;
      inSimulationMode : Bool;
      inStepStartTime : Int := 10;
      inStepEndTime : Int := 10;
   END_VAR
   VAR_OUTPUT
      outStepNb : Int;
      outStepStart : Bool;
   END_VAR
   VAR_IN_OUT
      inStepEnd : Bool;
      inManualStepNb : Int;
      inManualStepUp : Bool;
      inManualStepDown : Bool;
   END_VAR
   VAR
      sStepNb : Int;
      sStepNbOld : Int;
      sStepNbPrevious : Int;
      sStepStartTime : Time;
      sStepEndTime : Time;
      sStepStart : Bool;
      tonStepStart : TON_TIME;
      tonStepEnd : TON_TIME;
   END_VAR
   VAR_TEMP
      tIntToStartTime : DInt;
      tIntToEndTime : DInt;
   END_VAR
BEGIN
   IF #inStart THEN

       REGION Operating Mode

           IF #inManualMode THEN

               #sStepNb := #inManualStepNb;

               REGION Step +/- 1

                   IF #inManualStepUp THEN

                       #sStepNb := #inNexStepNb;

                   ELSIF #inManualStepDown THEN

                       #sStepNb := #sStepNbPrevious;

                   END_IF;

               END_REGION

           ELSE

                IF #sStepNb = 0 THEN

                    #sStepNb := 1;

               ELSIF #tonStepEnd.Q THEN

                   #sStepNb := #inNexStepNb;
                   #inStepEnd := FALSE;

               END_IF;

           END_IF;

       END_REGION

   ELSE

       #sStepNb := 0;
       #inStepEnd := FALSE;

   END_IF;

   REGION Step Start 

       IF #inStart AND #sStepNb<>#sStepNbOld OR NOT #inStart THEN

           #sStepStart := FALSE;
       ELSE

           #sStepStart := TRUE;

       END_IF;


   END_REGION


       REGION Rewriting time start/end step to timer

           //Czas poczatku i konca kroku zdefiniowany dla calej sekwencji
           //Mozna go nadpisywac w krokach 
           #tIntToStartTime := 1000 * #inStepStartTime;
           #tIntToEndTime := 1000 * #inStepEndTime;

           #sStepStartTime := DINT_TO_TIME(#tIntToStartTime);
           #sStepEndTime := DINT_TO_TIME(#tIntToEndTime);

       END_REGION

   REGION Step start/end delay timers

       REGION Step start timer

           #tonStepStart(IN := #sStepStart,
                         PT := #sStepStartTime);

       END_REGION

       REGION Step end timer

           #tonStepEnd(IN := #inStepEnd,
                       PT := #sStepEndTime);

       END_REGION

   END_REGION

   REGION Step old

       IF #sStepNb<>#sStepNbOld THEN

           #sStepNbPrevious := #sStepNbOld;

       END_IF;

       #sStepNbOld := #sStepNb;

   END_REGION

   REGION Reset impuls signals

       #inManualStepUp := FALSE;
       #inManualStepDown := FALSE;


   END_REGION

   REGION Outputs

       #inManualStepNb := #sStepNb;

       #outStepNb := #sStepNb;

       #outStepStart := #tonStepStart.Q AND NOT #inSimulationMode;

   END_REGION
END_FUNCTION_BLOCK

FUNCTION_BLOCK "Sequence1"   // FB5, SCL
{ S7_Optimized_Access := 'TRUE' }
VERSION : 0.1
   VAR
      Sequencer : "Sequencer";
      Static_1 : Bool;
   END_VAR
BEGIN

           #Sequencer.inStepStartTime := 2;
           #Sequencer.inStepEndTime := 2;

       CASE #Sequencer.outStepNb OF

           0: //Krok 0 Manual
               REGION Krok 0 Manual

                   #Sequencer.inNexStepNb := 1;

               END_REGION

           1:  // Krok 1
               REGION Krok 1

                   IF #Sequencer.outStepStart THEN
                       // DM Class activations

                       "DB_DM".pump2Tank1in.inTurnOn := TRUE;

                   END_IF;

                   // Next step 

                   IF "Tag_4" THEN

                       #Sequencer.inNexStepNb := 2;

                   ELSE

                       #Sequencer.inNexStepNb := 3;

                   END_IF;

                   // Step end

                   #Sequencer.inStepEnd := "Tag_5";

               END_REGION

               #Sequencer.inStepEndTime := 15;

           2:  // Krok 2

               REGION Krok 2

                   // DM Class activations

                   "DB_DM".pump2Tank1in.inTurnOn := TRUE;

               END_REGION

               // Step end

               #Sequencer.inStepEnd := "Tag_6";

               #Sequencer.inNexStepNb := 3;

          3: //Krok 3

              REGION Krok 3

                  // DM Class activations

                  "DB_DM".pump2Tank1in.inTurnOn := TRUE;


                  // DV Class activations

                  //ddd


                  // "PID" Setpoint

                  "PID_Tank1Level".Setpoint := 50;


                  // Sinamics Setpoint

                  "DB_Sinamics".pump2Control.Velocity := "PID_Tank1Level".Output;

                  "DB_Sinamics".pump1Control.Velocity := 100;

                  //

                  #Sequencer.inNexStepNb := 4;

                  #Sequencer.inStepEnd := "Tag_7";

              END_REGION

          4:  // Krok 4

              REGION Krok 4

                  // DM Class activations

                  "DB_DM".pump2Tank1in.inTurnOn := TRUE;

              END_REGION

              // Step end

              #Sequencer.inStepEnd := "Tag_6";

              #Sequencer.inStart := FALSE;

           ELSE  // Statement section ELSE

               #Sequencer.inStepEnd := FALSE;

       END_CASE;


       #Sequencer();
END_FUNCTION_BLOCK

FUNCTION "PID" : Void   // FC1, LAD
{ S7_Optimized_Access := 'TRUE' }
VERSION : 0.1
BEGIN

REGION Network 1
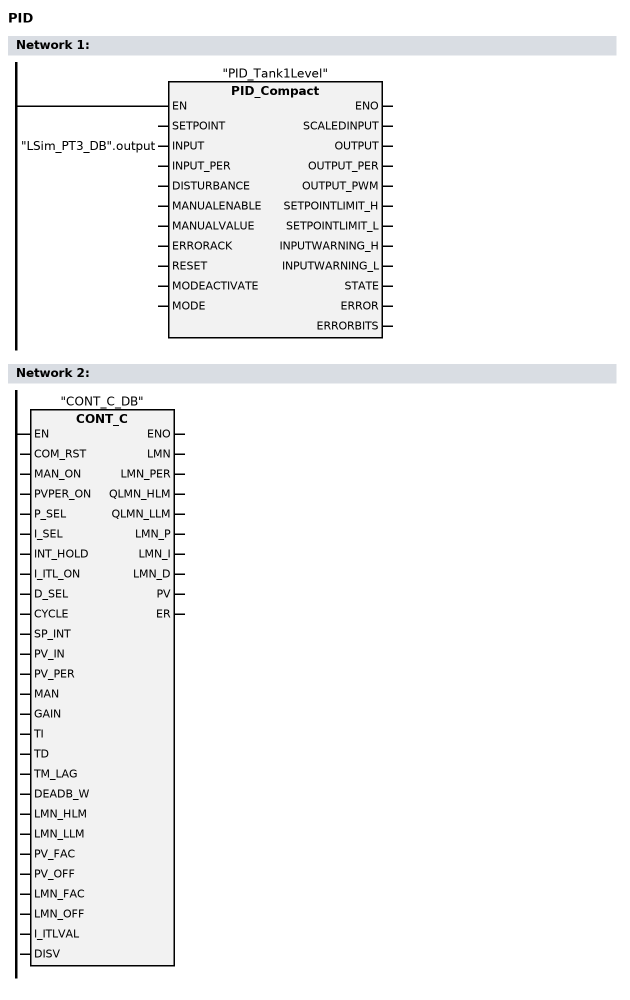
   "PID_Tank1Level"(Input := "LSim_PT3_DB".output);   // PID_Compact
END_REGION

REGION Network 2
   "CONT_C_DB"();   // CONT_C
END_REGION
END_FUNCTION

ORGANIZATION_BLOCK "Main"   // OB1, LAD, ProgramCycle
TITLE = "Main Program Sweep (Cycle)"
{ S7_Optimized_Access := 'TRUE' }
VERSION : 0.1
   VAR_INPUT
      Initial_Call : Bool;   // Initial call of this OB
      Remanence : Bool;   // =True, if remanent data are available
   END_VAR
BEGIN

REGION Network 1
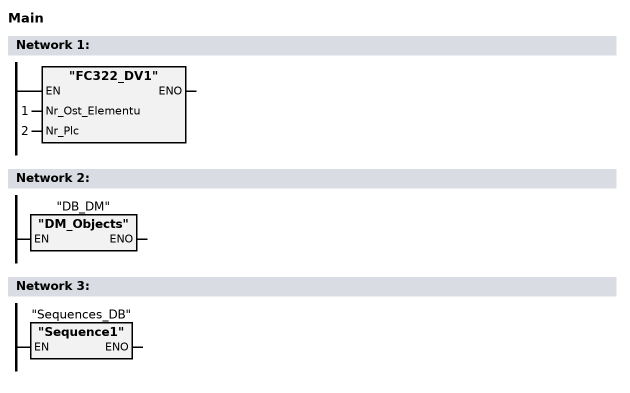
   RUNG wire#powerrail
      "FC322_DV1"(Nr_Ost_Elementu := 1, Nr_Plc := 2)
   END_RUNG
   // the same network as SCL:
   "FC322_DV1"(Nr_Ost_Elementu := 1, Nr_Plc := 2);
END_REGION

REGION Network 2
   RUNG wire#powerrail
      "DB_DM"()
   END_RUNG
   // the same network as SCL:
   "DB_DM"();   // "DM_Objects"
END_REGION

REGION Network 3
   RUNG wire#powerrail
      "Sequences_DB"()
   END_RUNG
   // the same network as SCL:
   "Sequences_DB"();   // "Sequence1"
END_REGION
END_ORGANIZATION_BLOCK

ORGANIZATION_BLOCK "Cyclic interrupt_20ms_PID"   // OB30, LAD, CyclicInterrupt
{ S7_Optimized_Access := 'TRUE' }
VERSION : 0.1
   VAR_INPUT
      Initial_Call : Bool;   // Initial call of this OB
      Event_Count : Int;   // Events discarded
   END_VAR
BEGIN

REGION Network 1
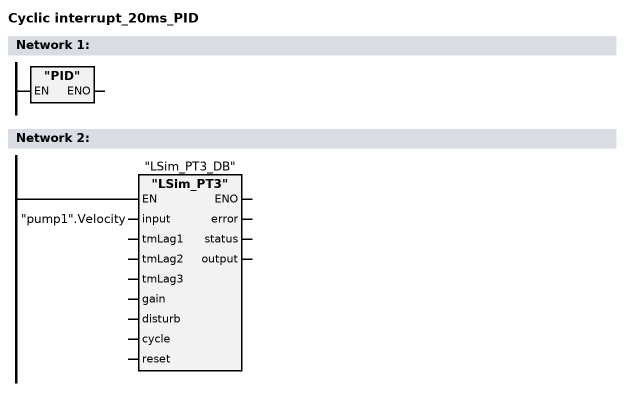
   RUNG wire#powerrail
      "PID"()
   END_RUNG
   // the same network as SCL:
   "PID"();
END_REGION

REGION Network 2
   RUNG wire#powerrail
      "LSim_PT3_DB"(input := "pump1".Velocity, tmLag1 :=, tmLag2 :=, tmLag3 :=, gain :=, disturb :=, cycle :=, reset :=, error =>, status =>, output =>)
   END_RUNG
   // the same network as SCL:
   "LSim_PT3_DB"(input := "pump1".Velocity);   // "LSim_PT3"
END_REGION
END_ORGANIZATION_BLOCK

ORGANIZATION_BLOCK "Cyclic interrupt_10ms_Sinamics"   // OB31, LAD, CyclicInterrupt
{ S7_Optimized_Access := 'TRUE' }
VERSION : 0.1
   VAR_INPUT
      Initial_Call : Bool;   // Initial call of this OB
      Event_Count : Int;   // Events discarded
   END_VAR
BEGIN

REGION Network 1
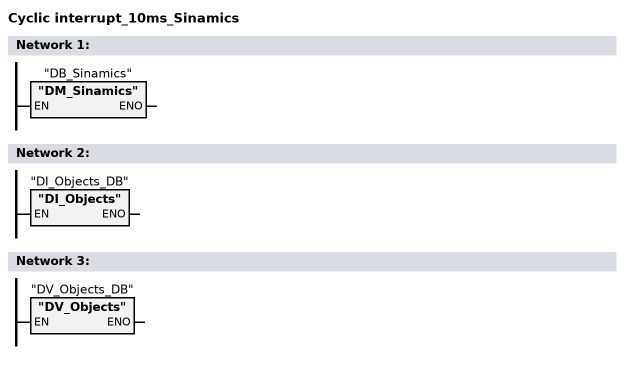
   RUNG wire#powerrail
      "DB_Sinamics"()
   END_RUNG
   // the same network as SCL:
   "DB_Sinamics"();   // "DM_Sinamics"
END_REGION

REGION Network 2
   RUNG wire#powerrail
      "DI_Objects_DB"()
   END_RUNG
   // the same network as SCL:
   "DI_Objects_DB"();   // "DI_Objects"
END_REGION

REGION Network 3
   RUNG wire#powerrail
      "DV_Objects_DB"()
   END_RUNG
   // the same network as SCL:
   "DV_Objects_DB"();   // "DV_Objects"
END_REGION
END_ORGANIZATION_BLOCK

// folder: DI

FUNCTION_BLOCK "DI_Objects"   // FB4, LAD
{ S7_Optimized_Access := 'TRUE' }
VERSION : 0.1
   VAR
      di1 : "DI_Class";
   END_VAR
BEGIN

REGION Network 2 (SCL)
   #di1();
END_REGION
END_FUNCTION_BLOCK

FUNCTION_BLOCK "DI_Class"   // FB300, SCL
{ S7_Optimized_Access := 'TRUE' }
VERSION : 0.1
   VAR_INPUT
      inActivateObject : Bool := true;   // Aktywowanie działania obiektu
      inLocalMode : Bool;   // Tryb lokalny
      inRemoteMode : Bool;   // Tryb remontowy
      inExtFault : Bool;   // Błąd zewnętrzny
      inLockAutoMan : Bool;   // Blokada przełączenia trybu Auto-Manual
      inInterlock : Bool;   // Interlok
      inGlobalAckFault : Bool;   // Globalny reset
      inAutoOff : Bool;   // Resetowanie sterowania na końcu
      inTurnOnDelay : DInt;   // Czas opóźnienia załączenia [s]
      inTurnOffDelay : DInt;   // Czas opóźnienia wyłączenia [s]
      inAlarmDelay : DInt;   // Czas opóźnienia alarmu od potwierdzeń [s]
   END_VAR
   VAR_OUTPUT
      oControl : Bool;   // Wyjście sterujące
      oAckFault : Bool;   // Wyjście reset obiektu
      oFault : Bool;   // Wyjście awaria
      oFaultCode : Byte;   // Kod awarii
      oStatusCode : Word;   // Kod statusu
      oStatus : Int;   // Status ( 1-awaria; 2-Wył; 4-Załączanie; 8-Zał; 16-Wyłączanie)
      oControlMode : Int;   // Tryb pracy (1-remont; 2-lokal; 4-manual; 8-auto)
   END_VAR
   VAR_IN_OUT
      inTurnOn : Bool;   // Załączanie z programu
      inCmdOper : Word := 16#5;   // Komendy manualne
      inSimOper : Word;   // Komendy symulacji
      inCmdOperImp : Word;   // Komendy impulsowe
   END_VAR
   VAR
      statManAuto : Bool;
      statSymOn : Bool;
      statSwitchEnable : Bool;
      statManTurnOn : Bool;
      statManDirection : Bool;
      statSwitchControl : Bool;
      statFaultReset : Bool;
      statActivate : Bool;
      statTurnOn : Bool;
      statLocal : Bool;
      statRemote : Bool;
      statExtFault : Bool;
      statLockAutoMan : Bool;
      statInterlock : Bool;
      tofTurnOnDelay : TON_TIME;
      tofTurnOffDelay : TOF_TIME;
      tonAlarm : TON_TIME;
      statAlarmStart : Bool;
      statFault : Bool;
      statControlMode : Int;
      statControl : Bool;
      statTmrOnOff : Bool;
      trigGlobalReset : R_TRIG;
   END_VAR
BEGIN
   REGION Activation object - condition to execute function
       IF NOT #inActivateObject THEN

           #inTurnOn := FALSE;
           #inCmdOper := 0;
           #inSimOper := 0;
           #inCmdOperImp := 0;

           #oControl := FALSE;
           #oAckFault := FALSE;
           #oFault := FALSE;
           #oFaultCode := 0;
           #oStatusCode := 0;
           #oStatus := 0;
           #oControlMode := 0;

           RETURN;

       END_IF;

   END_REGION

   REGION Rewriting inputs

       //Operator Control Word
       #statManAuto := #inCmdOper.%X0;
       #statSymOn := #inCmdOper.%X1;
       #statSwitchEnable := #inCmdOper.%X2;
       #statManTurnOn := #inCmdOper.%X3;
       #statManDirection := #inCmdOper.%X4;
       #statSwitchControl := #inCmdOper.%X6;

       //Operator Control Word Impulses
       #trigGlobalReset(CLK:=#inGlobalAckFault);

       #statFaultReset := #trigGlobalReset.Q OR #inCmdOperImp.%X0;

   END_REGION

   REGION Rewriting inputs or simulation signals to statics

       IF NOT #statSymOn THEN

           #statTurnOn := #inTurnOn;
           #statLocal := #inLocalMode;
           #statRemote := #inRemoteMode;
           #statExtFault := #inExtFault;
           #statLockAutoMan := #inLockAutoMan;
           #statInterlock := #inInterlock;

           //Rewriting inputs to simulation bits when simulotion is to switch fluently
           #inSimOper.%X0 := #statActivate;
           #inSimOper.%X1 := #statTurnOn;
           #inSimOper.%X5 := #statLocal;
           #inSimOper.%X6 := #statRemote;
           #inSimOper.%X7 := #statExtFault;
           #inSimOper.%X8 := #statLockAutoMan;
           #inSimOper.%X9 := #statInterlock;

       ELSE

           #statActivate := #inSimOper.%X0;
           #statTurnOn := #inSimOper.%X1;
           #statLocal := #inSimOper.%X5;
           #statRemote := #inSimOper.%X6;
           #statExtFault := #inSimOper.%X7;
           #statLockAutoMan := #inSimOper.%X8;
           #statInterlock := #inSimOper.%X9;

       END_IF;


   END_REGION

   REGION Control Mode

       IF #statRemote THEN

           #statControlMode := 1;

       ELSIF #statLocal THEN

           #statControlMode := 2;

       ELSIF NOT #statManAuto AND NOT #statLockAutoMan THEN

           #statControlMode := 4;

       ELSIF #statManAuto AND NOT #statLockAutoMan THEN

           #statControlMode := 8;

       END_IF;

   END_REGION

   REGION TurnOn/Off Delay

       #tofTurnOnDelay(IN := #statTurnOn,
                       PT := 1000 * #inTurnOnDelay);

       #tofTurnOffDelay(IN := #statTurnOn,
                        PT := 1000 * #inTurnOffDelay);

       IF #tofTurnOnDelay.Q THEN

           #statTmrOnOff := TRUE;

       END_IF;

       IF NOT #tofTurnOffDelay.Q THEN

           #statTmrOnOff := FALSE;

       END_IF;
   END_REGION

   REGION Fault 
       //Zerowanie czasu awari przy zmianie sterowanie podczas ruchu - czy to w ogole cokolwiek robi???



       //Generating fault
       IF #statExtFault THEN

           #statFault := TRUE;

       ELSIF #statFaultReset THEN

           #statFault := FALSE;

       END_IF;

       //Fault reset 
       // IF #statFaultReset THEN
       //     #statFault := FALSE;


       // END_IF;

       //Fault code
       #oFaultCode.%X2 := #statExtFault;

   END_REGION

   REGION Command locks

       IF #statControlMode = 8 AND #statLockAutoMan THEN

           #statManAuto := TRUE;

       ELSIF #statControlMode = 4 AND #statLockAutoMan THEN

           #statManAuto := FALSE;

       END_IF;

       // Writing states from Local to Manual when object when switching Local to Manual
       IF #statControlMode = 2 THEN

           #statManAuto := FALSE;

       END_IF;

       // Writing states from Auto to Manual when object when switching Auto to Manual
       // Przypadek gdy ktos z wlaczonym automatycznie urz. przechodzi na tryb zdalny-reczny
       IF #statControlMode = 8 THEN

           #statManTurnOn := #statTurnOn;

       END_IF;

       //Resetowanie rozkazu zalaczenia w trybie manualnym po awarii
       IF #statFault THEN

           #statManTurnOn := FALSE;

       END_IF;




   END_REGION

   REGION Control output

       #statControl :=
       #statSwitchEnable AND
       NOT #statInterlock AND
       NOT #statFault AND
       ((#statControlMode = 8 AND #statTmrOnOff) OR
       (#statControlMode = 4 AND #statManTurnOn));

   END_REGION

   REGION Reset Control

       #oAckFault := #statFaultReset;

   END_REGION ;

   REGION Device status code
       IF #statFault THEN
           #oStatus := 1;

       ELSIF #statControlMode = 1 THEN
           #oStatus := 2;

       ELSIF #statControlMode = 2 THEN

           IF #statControl THEN
               #oStatus := 4;

           ELSIF NOT #statControl THEN
               #oStatus := 16;
           END_IF;

       ELSIF #statControlMode > 2 THEN

           IF #statSwitchControl AND #statSwitchEnable THEN

               IF #statControl THEN

                   #oStatus := 4;

               ELSIF NOT #statControl THEN

                   #oStatus := 16;